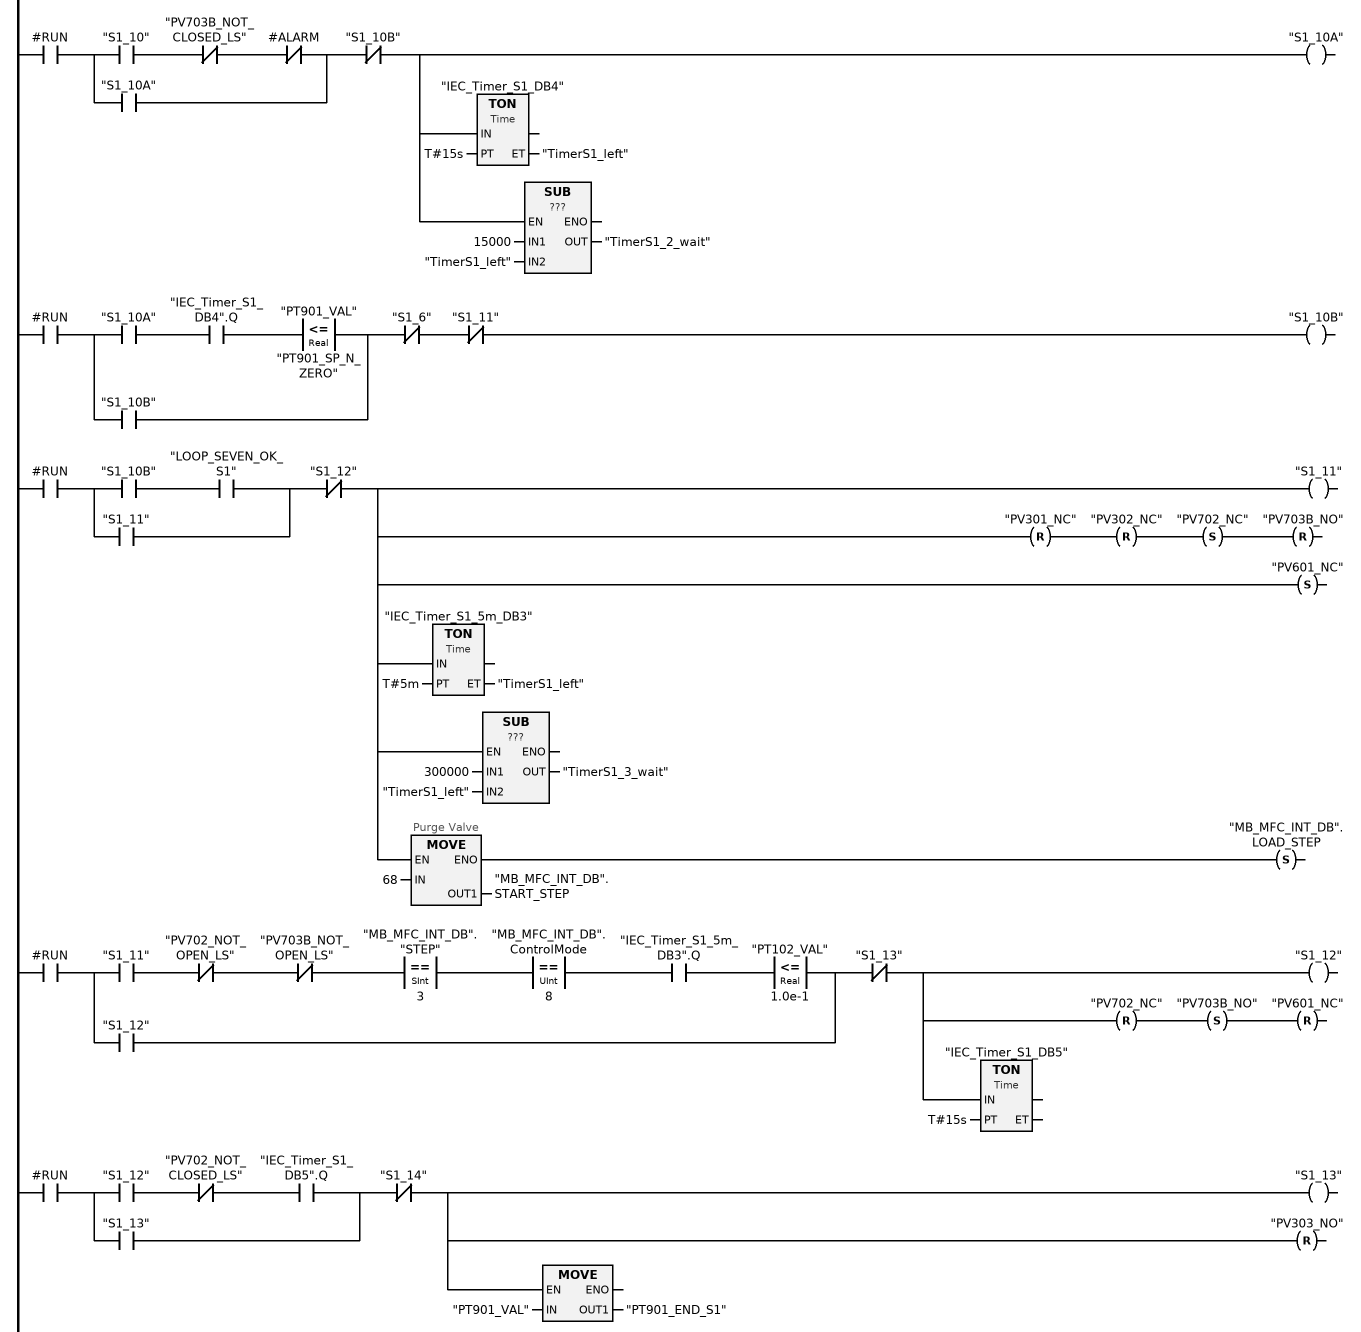
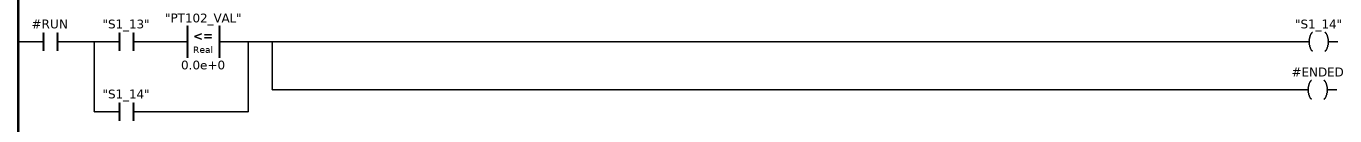
   "S1_0" := #RUN AND ((#START AND NOT #ALARM) OR "S1_0") AND NOT "S1_1";
   IF "S1_0" THEN
       "MB_MFC_INT_DB".MFC_MODE_SP := "MB_VAL_CONTROL_MODE_BUS";
       "MB_MFC_INT_DB".MFC_Setpoint := 0;
       "MB_MFC_INT_DB".START_STEP := 10;
       "MB_MFC_INT_DB".LOAD_STEP := TRUE;
       "MB_MFC_FLOAT_DB"."STEP" := -1;
   END_IF;
   "Timer_S1_DB_1S".TON(IN := "S1_0", PT := T#1S);
   IF "S1_0" THEN
       "GREEN_LIGHT" := FALSE;
       "YELLOW_LIGHT" := TRUE;
   END_IF;
   "S1_1" := #RUN AND (("S1_0" AND "Timer_S1_DB_1S".Q AND ("MB_MFC_INT_DB"."STEP" = 3) AND NOT #ALARM) OR "S1_1") AND NOT "S1_1A";
   IF "S1_1" THEN "PV703A_NO" := FALSE; END_IF;
   "S1_1A" := #RUN AND (("S1_1" AND NOT "PV703A_NOT_OPEN_LS" AND NOT #ALARM) OR "S1_1A") AND NOT "S1_2";
   IF "S1_1A" THEN
       "PV303_NO" := TRUE;
       "PV301_NC" := TRUE;
       "PV302_NC" := TRUE;
       "MB_MFC_INT_DB".MFC_Setpoint := "STEP1_MFC_FL_SP";
       "MB_MFC_INT_DB".START_STEP := 10;
       "MB_MFC_INT_DB".LOAD_STEP := TRUE;
   END_IF;
   "S1_2" := #RUN AND (("S1_1A" AND NOT #ALARM AND ("PT302_VAL" < "PT302_HIGH") AND ("MB_MFC_INT_DB"."STEP" = 3) AND ("MB_MFC_INT_DB".MFC_Setpoint = "STEP1_MFC_FL_SP")) OR "S1_2") AND NOT "S1_3";
   IF "S1_2" THEN "PV601_NC" := TRUE; END_IF;
   "S1_3" := #RUN AND (("S1_2" AND NOT #ALARM AND ("PT601_VAL" >= "PT302_CALC_90PRCT")) OR "S1_3") AND NOT "S1_4";
   IF "S1_3" THEN "PV702_NC" := TRUE; END_IF;
   "Timer_S1_DB_3S".TON(IN := "S1_3", PT := T#1.5s, ET => "TempDWord_A");
   "S1_4" := #RUN AND (("S1_3" AND "Timer_S1_DB_3S".Q AND NOT "PV702_NOT_OPEN_LS" AND NOT #ALARM) OR "S1_4") AND NOT "S1_5";
   IF "S1_4" THEN
       "PV601_NC" := FALSE;
       "PV702_NC" := FALSE;
   END_IF;
   "S1_5" := #RUN AND (("S1_4" AND NOT "PV702_NOT_CLOSED_LS" AND NOT #ALARM) OR "S1_5") AND NOT "S1_6";
   "IEC_Counter_S1_1".CTU(CU := "S1_7", R := "S1_2", PV := "STEP1_LOOPS", CV => "Counter_S1");
   "LOOP_SEVEN_OK_S1" := "IEC_Counter_S1_1".Q;
   "S1_6" := #RUN AND ((("S1_5" OR ("S1_10B" AND NOT "LOOP_SEVEN_OK_S1")) AND NOT #ALARM) OR "S1_6") AND NOT "S1_7";
   IF "S1_6" THEN
       "PV701_NC" := TRUE;
       "PT901_SAVE" := "PT901_VAL" - 1.0;
   END_IF;
   IF "S1_6" AND ("PT601_VAL" < 3.5) THEN "PV601_NC" := TRUE; END_IF;
   "S1_7" := #RUN AND (("S1_6" AND NOT "PV701_NOT_OPEN_LS" AND ("PT901_VAL" >= "PT901_SP_N")) OR "S1_7") AND NOT "S1_7A";
   IF "S1_7" THEN
       "PV701_NC" := FALSE;
       "PV601_NC" := FALSE;
   END_IF;
   "S1_7A" := #RUN AND (("S1_7" AND NOT "PV701_NOT_CLOSED_LS" AND "Timer_S1_DB_5S".Q AND ("PT901_VAL" >= "PT901_SAVE")) OR "S1_7A") AND NOT "S1_8";
   "S1_8" := #RUN AND (("S1_7A" AND NOT #ALARM) OR "S1_8") AND NOT "S1_9";
   IF "S1_8" THEN "PV703B_NO" := FALSE; END_IF;
   "S1_9" := #RUN AND (("S1_8" AND NOT "PV703B_NOT_OPEN_LS" AND ("PT901_VAL" <= "PT901_SP_PV703B_OPEN") AND NOT #ALARM) OR "S1_9") AND NOT "S1_10";
   "IEC_Timer_S1_DB3".TON(IN := "S1_9", PT := T#150s, ET => "TimerS1_left");
   IF "S1_9" THEN "TimerS1_1_wait" := 150000 - "TimerS1_left"; END_IF;
   "S1_10" := #RUN AND (("S1_9" AND "IEC_Timer_S1_DB3".Q AND ("PT901_VAL" <= 0.2)) OR "S1_10") AND NOT "S1_10A";
   IF "S1_10" THEN "PV703B_NO" := TRUE; END_IF;
   "S1_10A" := #RUN AND (("S1_10" AND NOT "PV703B_NOT_CLOSED_LS" AND NOT #ALARM) OR "S1_10A") AND NOT "S1_10B";
   "IEC_Timer_S1_DB4".TON(IN := "S1_10A", PT := T#15s, ET => "TimerS1_left");
   IF "S1_10A" THEN "TimerS1_2_wait" := 15000 - "TimerS1_left"; END_IF;
   "S1_10B" := #RUN AND (("S1_10A" AND "IEC_Timer_S1_DB4".Q AND ("PT901_VAL" <= "PT901_SP_N_ZERO")) OR "S1_10B") AND NOT "S1_6" AND NOT "S1_11";
   "S1_11" := #RUN AND (("S1_10B" AND "LOOP_SEVEN_OK_S1") OR "S1_11") AND NOT "S1_12";
   IF "S1_11" THEN
       "PV301_NC" := FALSE;
       "PV302_NC" := FALSE;
       "PV702_NC" := TRUE;
       "PV703B_NO" := FALSE;
       "PV601_NC" := TRUE;
   END_IF;
   "IEC_Timer_S1_5m_DB3".TON(IN := "S1_11", PT := T#5m, ET => "TimerS1_left");
   IF "S1_11" THEN
       "TimerS1_3_wait" := 300000 - "TimerS1_left";
       "MB_MFC_INT_DB".START_STEP := 68;   // Purge Valve
       "MB_MFC_INT_DB".LOAD_STEP := TRUE;
   END_IF;
   "S1_12" := #RUN AND (("S1_11" AND NOT "PV702_NOT_OPEN_LS" AND NOT "PV703B_NOT_OPEN_LS" AND ("MB_MFC_INT_DB"."STEP" = 3) AND ("MB_MFC_INT_DB".ControlMode = 8) AND "IEC_Timer_S1_5m_DB3".Q AND ("PT102_VAL" <= 1.0e-1)) OR "S1_12") AND NOT "S1_13";
   IF "S1_12" THEN
       "PV702_NC" := FALSE;
       "PV703B_NO" := TRUE;
       "PV601_NC" := FALSE;
   END_IF;
   "IEC_Timer_S1_DB5".TON(IN := "S1_12", PT := T#15s);
   "S1_13" := #RUN AND (("S1_12" AND NOT "PV702_NOT_CLOSED_LS" AND "IEC_Timer_S1_DB5".Q) OR "S1_13") AND NOT "S1_14";
   IF "S1_13" THEN
       "PV303_NO" := FALSE;
       "PT901_END_S1" := "PT901_VAL";
   END_IF;
   "S1_14" := #RUN AND (("S1_13" AND ("PT102_VAL" <= 0.0e+0)) OR "S1_14");
   #ENDED := "S1_14";
END_REGION

REGION Network 4
   // Timers
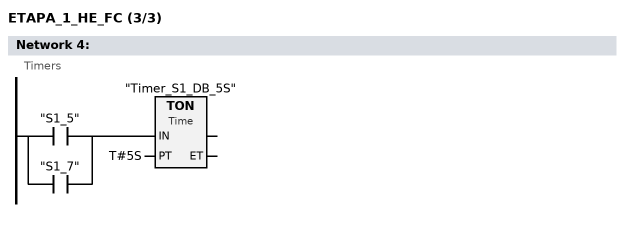
   "Timer_S1_DB_5S".TON(IN := "S1_5" OR "S1_7", PT := T#5S);
END_REGION
END_FUNCTION

FUNCTION "MB_READ_MX" : Void   // FC23, LAD
{ S7_Optimized_Access := 'FALSE' }
VERSION : 0.1
   VAR_TEMP   // added for the SCL form of the ladder/FBD networks
      _w1 : Bool;
      _w2 : Bool;
   END_VAR
BEGIN

REGION Network 1
   // MODBUS MASTER Cyclic Read
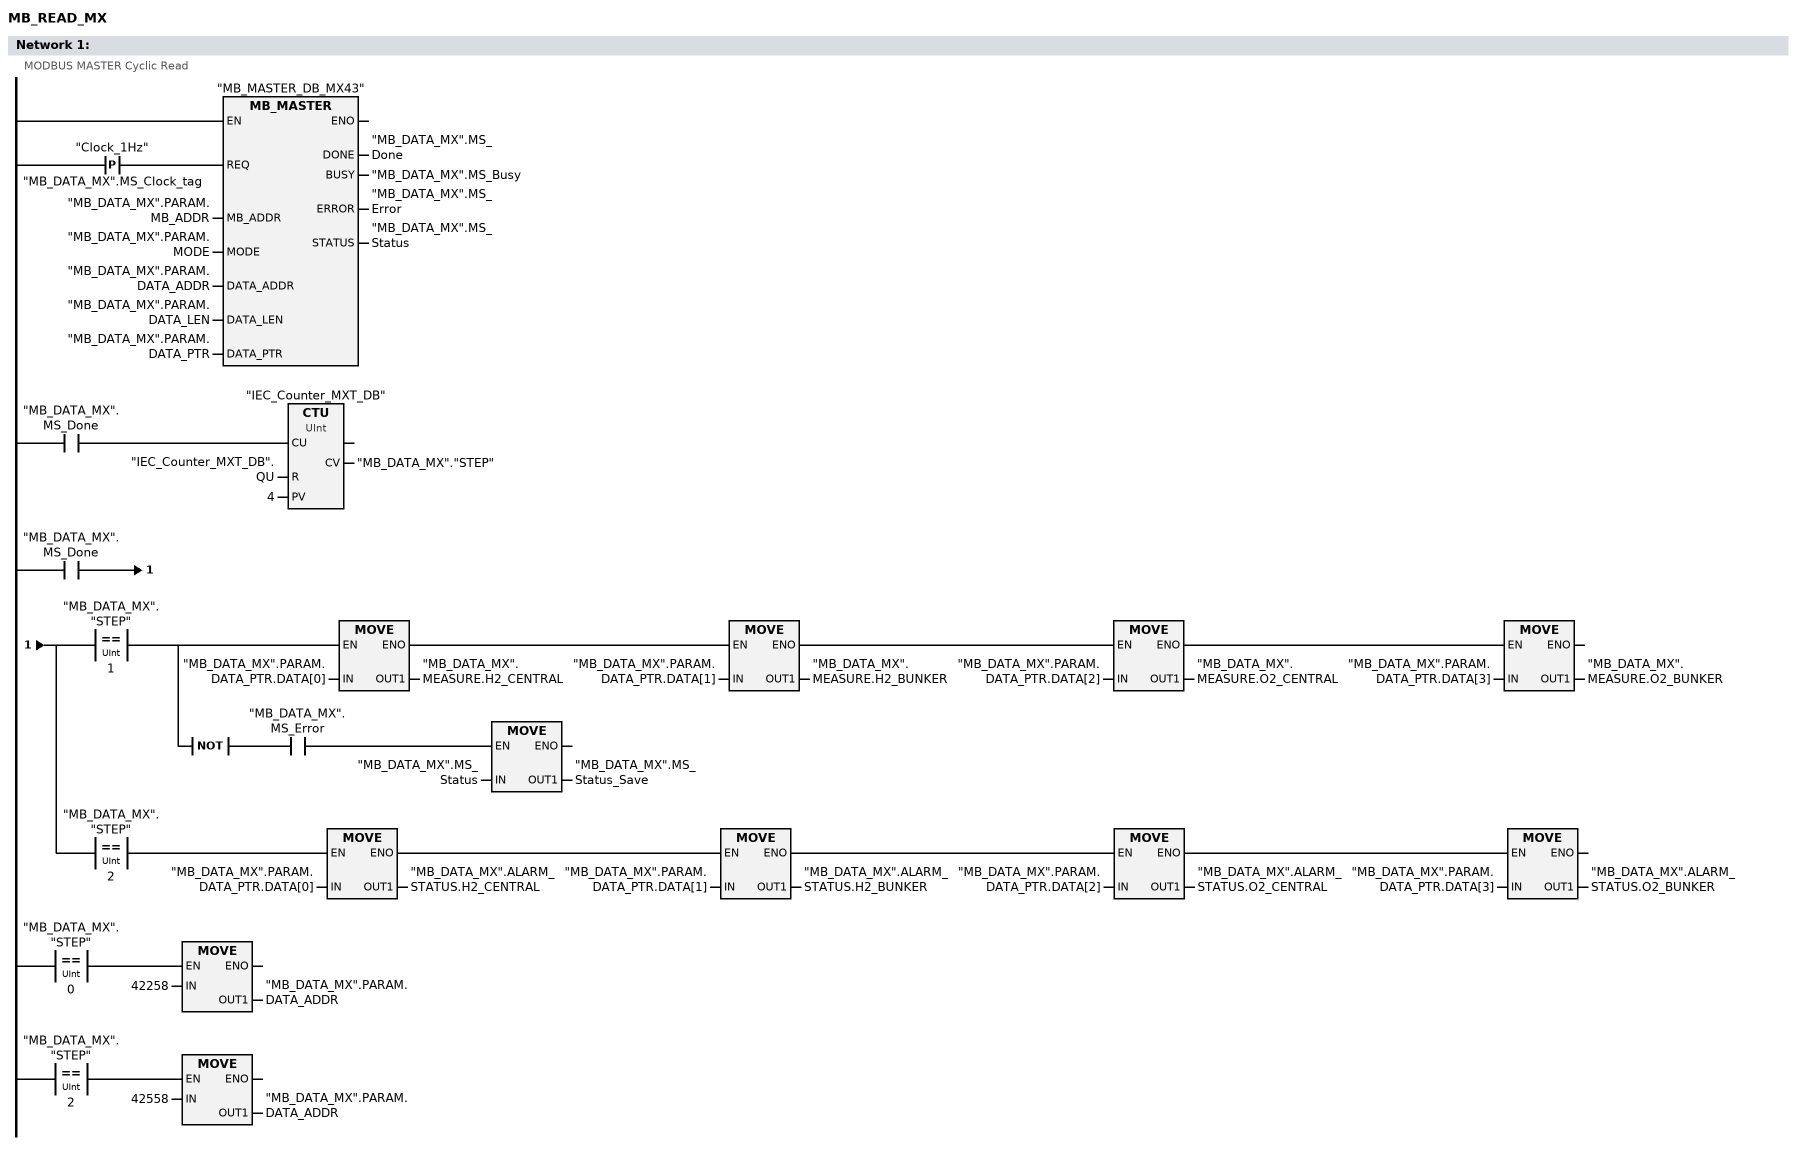
   #_w1 := "Clock_1Hz" AND NOT "MB_DATA_MX".MS_Clock_tag;   // rising edge of "Clock_1Hz"
   "MB_DATA_MX".MS_Clock_tag := "Clock_1Hz";
   "MB_MASTER_DB_MX43"(REQ := #_w1,   // MB_MASTER
                       MB_ADDR := "MB_DATA_MX".PARAM.MB_ADDR,
                       MODE := "MB_DATA_MX".PARAM.MODE,
                       DATA_ADDR := "MB_DATA_MX".PARAM.DATA_ADDR,
                       DATA_LEN := "MB_DATA_MX".PARAM.DATA_LEN,
                       DATA_PTR := "MB_DATA_MX".PARAM.DATA_PTR,
                       DONE => "MB_DATA_MX".MS_Done,
                       BUSY => "MB_DATA_MX".MS_Busy,
                       ERROR => "MB_DATA_MX".MS_Error,
                       STATUS => "MB_DATA_MX".MS_Status);
   "IEC_Counter_MXT_DB".CTU(CU := "MB_DATA_MX".MS_Done,
                           R := "IEC_Counter_MXT_DB".QU,
                           PV := 4,
                           CV => "MB_DATA_MX"."STEP");
   #_w2 := "MB_DATA_MX".MS_Done AND ("MB_DATA_MX"."STEP" = 1);
   IF #_w2 THEN
       "MB_DATA_MX".MEASURE.H2_CENTRAL := "MB_DATA_MX".PARAM.DATA_PTR.DATA[0];
       "MB_DATA_MX".MEASURE.H2_BUNKER := "MB_DATA_MX".PARAM.DATA_PTR.DATA[1];
       "MB_DATA_MX".MEASURE.O2_CENTRAL := "MB_DATA_MX".PARAM.DATA_PTR.DATA[2];
       "MB_DATA_MX".MEASURE.O2_BUNKER := "MB_DATA_MX".PARAM.DATA_PTR.DATA[3];
   END_IF;
   IF NOT #_w2 AND "MB_DATA_MX".MS_Error THEN "MB_DATA_MX".MS_Status_Save := "MB_DATA_MX".MS_Status; END_IF;
   IF "MB_DATA_MX".MS_Done AND ("MB_DATA_MX"."STEP" = 2) THEN
       "MB_DATA_MX".ALARM_STATUS.H2_CENTRAL := "MB_DATA_MX".PARAM.DATA_PTR.DATA[0];
       "MB_DATA_MX".ALARM_STATUS.H2_BUNKER := "MB_DATA_MX".PARAM.DATA_PTR.DATA[1];
       "MB_DATA_MX".ALARM_STATUS.O2_CENTRAL := "MB_DATA_MX".PARAM.DATA_PTR.DATA[2];
       "MB_DATA_MX".ALARM_STATUS.O2_BUNKER := "MB_DATA_MX".PARAM.DATA_PTR.DATA[3];
   END_IF;
   IF "MB_DATA_MX"."STEP" = 0 THEN "MB_DATA_MX".PARAM.DATA_ADDR := 42258; END_IF;
   IF "MB_DATA_MX"."STEP" = 2 THEN "MB_DATA_MX".PARAM.DATA_ADDR := 42558; END_IF;
END_REGION
END_FUNCTION

ORGANIZATION_BLOCK "Main"   // OB1, LAD, ProgramCycle
TITLE = "Main Program Sweep (Cycle)"
{ S7_Optimized_Access := 'FALSE' }
VERSION : 0.1
// Main with He Purging, Step 2 is Bypassed
   VAR_TEMP   // added for the SCL form of the ladder/FBD networks
      _w1 : Bool;
   END_VAR
BEGIN

REGION Network 1
   // TOP LOGIC
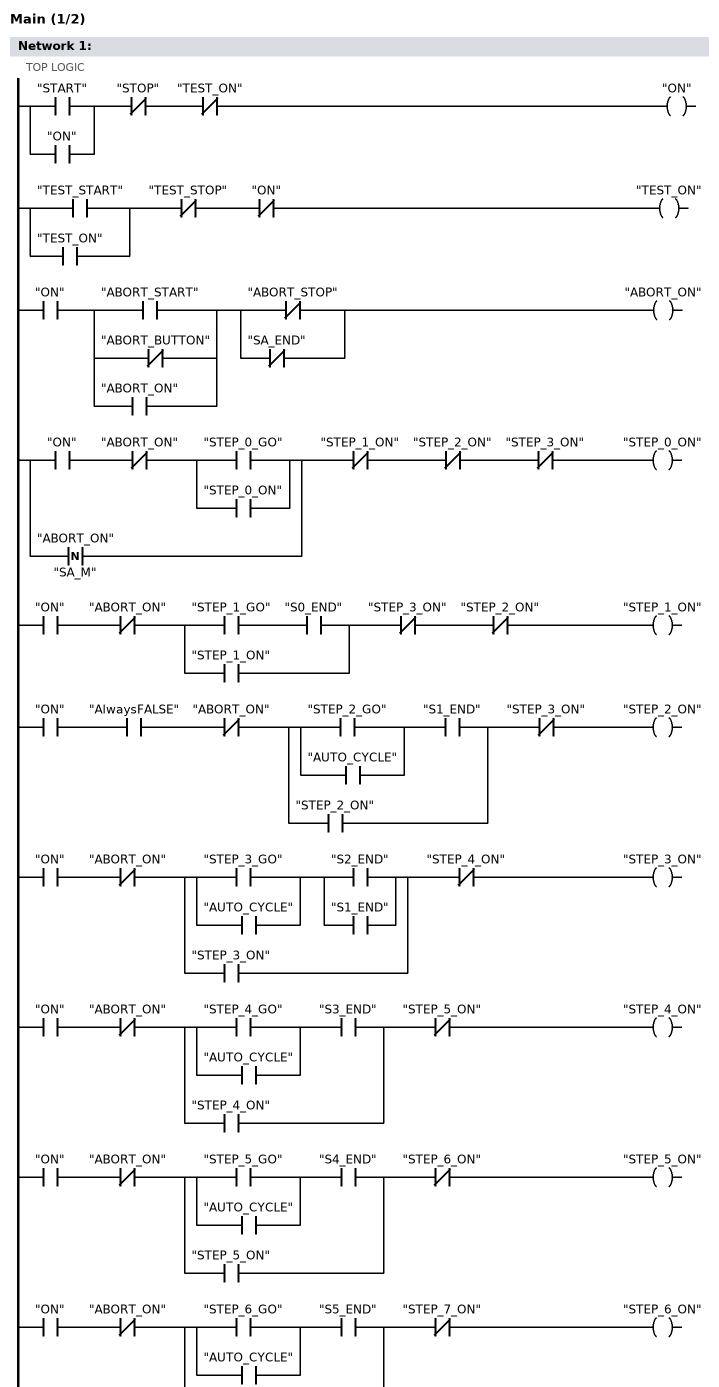
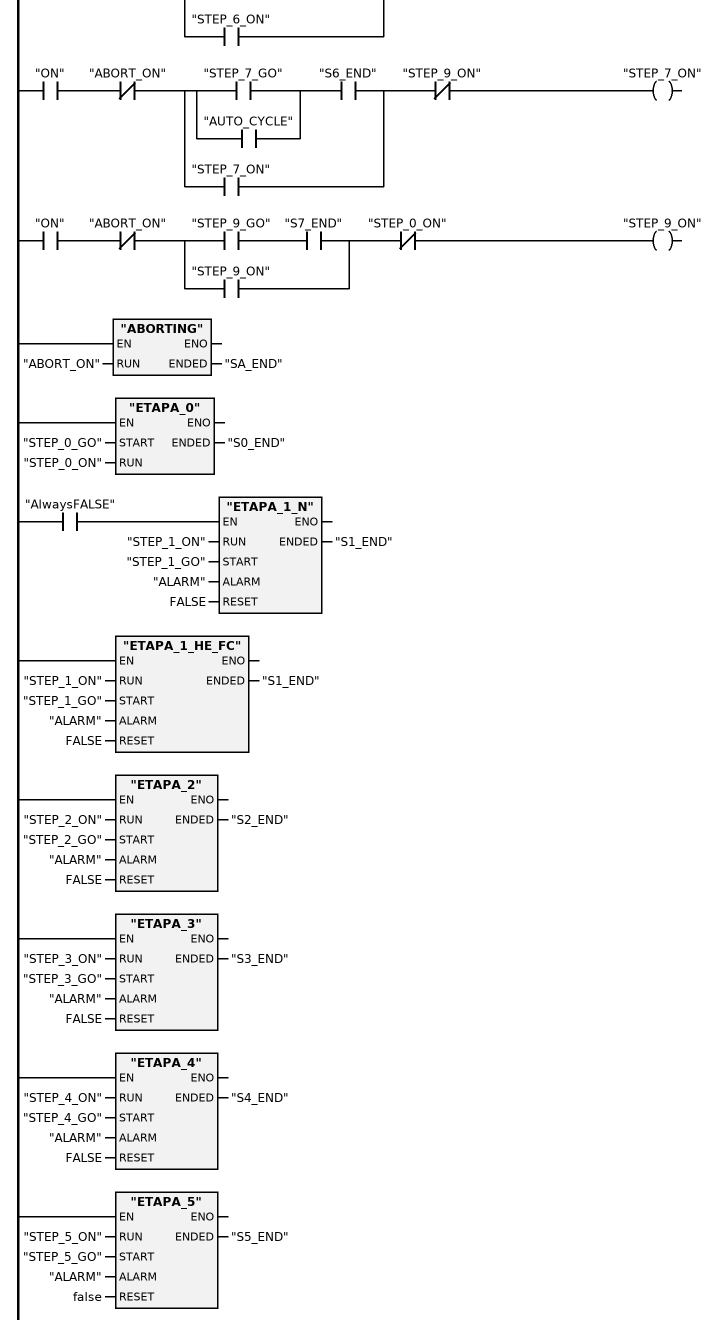
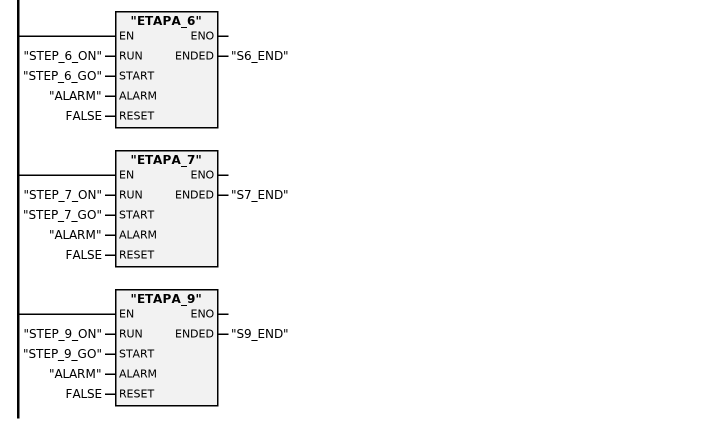
   RUNG wire#powerrail
      Contact( "START" )
      wire#w1
      I_Contact( "STOP" )
      I_Contact( "TEST_ON" )
      Coil( "ON" )
   END_RUNG
   RUNG wire#powerrail
      Contact( "ON" )
   END_RUNG wire#w1
   RUNG wire#powerrail
      Contact( "TEST_START" )
      wire#w2
      I_Contact( "TEST_STOP" )
      I_Contact( "ON" )
      Coil( "TEST_ON" )
   END_RUNG
   RUNG wire#powerrail
      Contact( "TEST_ON" )
   END_RUNG wire#w2
   RUNG wire#powerrail
      Contact( "ON" )
      wire#w3
      Contact( "ABORT_START" )
      wire#w4
      I_Contact( "ABORT_STOP" )
      wire#w5
      Coil( "ABORT_ON" )
   END_RUNG
   RUNG wire#w3
      I_Contact( "ABORT_BUTTON" )
   END_RUNG wire#w4
   RUNG wire#w3
      Contact( "ABORT_ON" )
   END_RUNG wire#w4
   RUNG wire#w4
      I_Contact( "SA_END" )
   END_RUNG wire#w5
   RUNG wire#powerrail
      Contact( "ON" )
      I_Contact( "ABORT_ON" )
      wire#w6
      Contact( "STEP_0_GO" )
      wire#w7
      I_Contact( "STEP_1_ON" )
      I_Contact( "STEP_2_ON" )
      I_Contact( "STEP_3_ON" )
      Coil( "STEP_0_ON" )
   END_RUNG
   RUNG wire#w6
      Contact( "STEP_0_ON" )
   END_RUNG wire#w7
   RUNG wire#powerrail
      N_Contact(operand := "ABORT_ON", bit := "SA_M")
   END_RUNG wire#w7
   RUNG wire#powerrail
      Contact( "ON" )
      I_Contact( "ABORT_ON" )
      wire#w8
      Contact( "STEP_1_GO" )
      Contact( "S0_END" )
      wire#w9
      I_Contact( "STEP_3_ON" )
      I_Contact( "STEP_2_ON" )
      Coil( "STEP_1_ON" )
   END_RUNG
   RUNG wire#w8
      Contact( "STEP_1_ON" )
   END_RUNG wire#w9
   RUNG wire#powerrail
      Contact( "ON" )
      Contact( "AlwaysFALSE" )
      I_Contact( "ABORT_ON" )
      wire#w10
      Contact( "STEP_2_GO" )
      wire#w11
      Contact( "S1_END" )
      wire#w12
      I_Contact( "STEP_3_ON" )
      Coil( "STEP_2_ON" )
   END_RUNG
   RUNG wire#w10
      Contact( "AUTO_CYCLE" )
   END_RUNG wire#w11
   RUNG wire#w10
      Contact( "STEP_2_ON" )
   END_RUNG wire#w12
   RUNG wire#powerrail
      Contact( "ON" )
      I_Contact( "ABORT_ON" )
      wire#w13
      Contact( "STEP_3_GO" )
      wire#w14
      Contact( "S2_END" )
      wire#w15
      I_Contact( "STEP_4_ON" )
      Coil( "STEP_3_ON" )
   END_RUNG
   RUNG wire#w13
      Contact( "AUTO_CYCLE" )
   END_RUNG wire#w14
   RUNG wire#w14
      Contact( "S1_END" )
   END_RUNG wire#w15
   RUNG wire#w13
      Contact( "STEP_3_ON" )
   END_RUNG wire#w15
   RUNG wire#powerrail
      Contact( "ON" )
      I_Contact( "ABORT_ON" )
      wire#w16
      Contact( "STEP_4_GO" )
      wire#w17
      Contact( "S3_END" )
      wire#w18
      I_Contact( "STEP_5_ON" )
      Coil( "STEP_4_ON" )
   END_RUNG
   RUNG wire#w16
      Contact( "AUTO_CYCLE" )
   END_RUNG wire#w17
   RUNG wire#w16
      Contact( "STEP_4_ON" )
   END_RUNG wire#w18
   RUNG wire#powerrail
      Contact( "ON" )
      I_Contact( "ABORT_ON" )
      wire#w19
      Contact( "STEP_5_GO" )
      wire#w20
      Contact( "S4_END" )
      wire#w21
      I_Contact( "STEP_6_ON" )
      Coil( "STEP_5_ON" )
   END_RUNG
   RUNG wire#w19
      Contact( "AUTO_CYCLE" )
   END_RUNG wire#w20
   RUNG wire#w19
      Contact( "STEP_5_ON" )
   END_RUNG wire#w21
   RUNG wire#powerrail
      Contact( "ON" )
      I_Contact( "ABORT_ON" )
      wire#w22
      Contact( "STEP_6_GO" )
      wire#w23
      Contact( "S5_END" )
      wire#w24
      I_Contact( "STEP_7_ON" )
      Coil( "STEP_6_ON" )
   END_RUNG
   RUNG wire#w22
      Contact( "AUTO_CYCLE" )
   END_RUNG wire#w23
   RUNG wire#w22
      Contact( "STEP_6_ON" )
   END_RUNG wire#w24
   RUNG wire#powerrail
      Contact( "ON" )
      I_Contact( "ABORT_ON" )
      wire#w25
      Contact( "STEP_7_GO" )
      wire#w26
      Contact( "S6_END" )
      wire#w27
      I_Contact( "STEP_9_ON" )
      Coil( "STEP_7_ON" )
   END_RUNG
   RUNG wire#w25
      Contact( "AUTO_CYCLE" )
   END_RUNG wire#w26
   RUNG wire#w25
      Contact( "STEP_7_ON" )
   END_RUNG wire#w27
   RUNG wire#powerrail
      Contact( "ON" )
      I_Contact( "ABORT_ON" )
      wire#w28
      Contact( "STEP_9_GO" )
      Contact( "S7_END" )
      wire#w29
      I_Contact( "STEP_0_ON" )
      Coil( "STEP_9_ON" )
   END_RUNG
   RUNG wire#w28
      Contact( "STEP_9_ON" )
   END_RUNG wire#w29
   RUNG wire#powerrail
      "ABORTING"(RUN := "ABORT_ON", ENDED => "SA_END")
   END_RUNG
   RUNG wire#powerrail
      "ETAPA_0"(START := "STEP_0_GO", RUN := "STEP_0_ON", ENDED => "S0_END")
   END_RUNG
   RUNG wire#powerrail
      Contact( "AlwaysFALSE" )
      "ETAPA_1_N"(RUN := "STEP_1_ON", START := "STEP_1_GO", ALARM := "ALARM", RESET := FALSE, ENDED => "S1_END")
   END_RUNG
   RUNG wire#powerrail
      "ETAPA_1_HE_FC"(RUN := "STEP_1_ON", START := "STEP_1_GO", ALARM := "ALARM", RESET := FALSE, ENDED => "S1_END")
   END_RUNG
   RUNG wire#powerrail
      "ETAPA_2"(RUN := "STEP_2_ON", START := "STEP_2_GO", ALARM := "ALARM", RESET := FALSE, ENDED => "S2_END")
   END_RUNG
   RUNG wire#powerrail
      "ETAPA_3"(RUN := "STEP_3_ON", START := "STEP_3_GO", ALARM := "ALARM", RESET := FALSE, ENDED => "S3_END")
   END_RUNG
   RUNG wire#powerrail
      "ETAPA_4"(RUN := "STEP_4_ON", START := "STEP_4_GO", ALARM := "ALARM", RESET := FALSE, ENDED => "S4_END")
   END_RUNG
   RUNG wire#powerrail
      "ETAPA_5"(RUN := "STEP_5_ON", START := "STEP_5_GO", ALARM := "ALARM", RESET := false, ENDED => "S5_END")
   END_RUNG
   RUNG wire#powerrail
      "ETAPA_6"(RUN := "STEP_6_ON", START := "STEP_6_GO", ALARM := "ALARM", RESET := FALSE, ENDED => "S6_END")
   END_RUNG
   RUNG wire#powerrail
      "ETAPA_7"(RUN := "STEP_7_ON", START := "STEP_7_GO", ALARM := "ALARM", RESET := FALSE, ENDED => "S7_END")
   END_RUNG
   RUNG wire#powerrail
      "ETAPA_9"(RUN := "STEP_9_ON", START := "STEP_9_GO", ALARM := "ALARM", RESET := FALSE, ENDED => "S9_END")
   END_RUNG
   // the same network as SCL:
   "ON" := ("START" OR "ON") AND NOT "STOP" AND NOT "TEST_ON";
   "TEST_ON" := ("TEST_START" OR "TEST_ON") AND NOT "TEST_STOP" AND NOT "ON";
   "ABORT_ON" := "ON" AND ("ABORT_START" OR NOT "ABORT_BUTTON" OR "ABORT_ON") AND (NOT "ABORT_STOP" OR NOT "SA_END");
   #_w1 := NOT "ABORT_ON" AND "SA_M";   // falling edge of "ABORT_ON"
   "SA_M" := "ABORT_ON";
   "STEP_0_ON" := (("ON" AND NOT "ABORT_ON" AND ("STEP_0_GO" OR "STEP_0_ON")) OR #_w1) AND NOT "STEP_1_ON" AND NOT "STEP_2_ON" AND NOT "STEP_3_ON";
   "STEP_1_ON" := "ON" AND NOT "ABORT_ON" AND (("STEP_1_GO" AND "S0_END") OR "STEP_1_ON") AND NOT "STEP_3_ON" AND NOT "STEP_2_ON";
   "STEP_2_ON" := "ON" AND "AlwaysFALSE" AND NOT "ABORT_ON" AND ((("STEP_2_GO" OR "AUTO_CYCLE") AND "S1_END") OR "STEP_2_ON") AND NOT "STEP_3_ON";
   "STEP_3_ON" := "ON" AND NOT "ABORT_ON" AND ((("STEP_3_GO" OR "AUTO_CYCLE") AND ("S2_END" OR "S1_END")) OR "STEP_3_ON") AND NOT "STEP_4_ON";
   "STEP_4_ON" := "ON" AND NOT "ABORT_ON" AND ((("STEP_4_GO" OR "AUTO_CYCLE") AND "S3_END") OR "STEP_4_ON") AND NOT "STEP_5_ON";
   "STEP_5_ON" := "ON" AND NOT "ABORT_ON" AND ((("STEP_5_GO" OR "AUTO_CYCLE") AND "S4_END") OR "STEP_5_ON") AND NOT "STEP_6_ON";
   "STEP_6_ON" := "ON" AND NOT "ABORT_ON" AND ((("STEP_6_GO" OR "AUTO_CYCLE") AND "S5_END") OR "STEP_6_ON") AND NOT "STEP_7_ON";
   "STEP_7_ON" := "ON" AND NOT "ABORT_ON" AND ((("STEP_7_GO" OR "AUTO_CYCLE") AND "S6_END") OR "STEP_7_ON") AND NOT "STEP_9_ON";
   "STEP_9_ON" := "ON" AND NOT "ABORT_ON" AND (("STEP_9_GO" AND "S7_END") OR "STEP_9_ON") AND NOT "STEP_0_ON";
   "ABORTING"(RUN := "ABORT_ON", ENDED => "SA_END");
   "ETAPA_0"(START := "STEP_0_GO", RUN := "STEP_0_ON", ENDED => "S0_END");
   IF "AlwaysFALSE" THEN
       "ETAPA_1_N"(RUN := "STEP_1_ON", START := "STEP_1_GO", ALARM := "ALARM", RESET := FALSE, ENDED => "S1_END");
   END_IF;
   "ETAPA_1_HE_FC"(RUN := "STEP_1_ON",
                   START := "STEP_1_GO",
                   ALARM := "ALARM",
                   RESET := FALSE,
                   ENDED => "S1_END");
   "ETAPA_2"(RUN := "STEP_2_ON", START := "STEP_2_GO", ALARM := "ALARM", RESET := FALSE, ENDED => "S2_END");
   "ETAPA_3"(RUN := "STEP_3_ON", START := "STEP_3_GO", ALARM := "ALARM", RESET := FALSE, ENDED => "S3_END");
   "ETAPA_4"(RUN := "STEP_4_ON", START := "STEP_4_GO", ALARM := "ALARM", RESET := FALSE, ENDED => "S4_END");
   "ETAPA_5"(RUN := "STEP_5_ON", START := "STEP_5_GO", ALARM := "ALARM", RESET := false, ENDED => "S5_END");
   "ETAPA_6"(RUN := "STEP_6_ON", START := "STEP_6_GO", ALARM := "ALARM", RESET := FALSE, ENDED => "S6_END");
   "ETAPA_7"(RUN := "STEP_7_ON", START := "STEP_7_GO", ALARM := "ALARM", RESET := FALSE, ENDED => "S7_END");
   "ETAPA_9"(RUN := "STEP_9_ON", START := "STEP_9_GO", ALARM := "ALARM", RESET := FALSE, ENDED => "S9_END");
END_REGION

REGION Network 2
   // ALARM Block
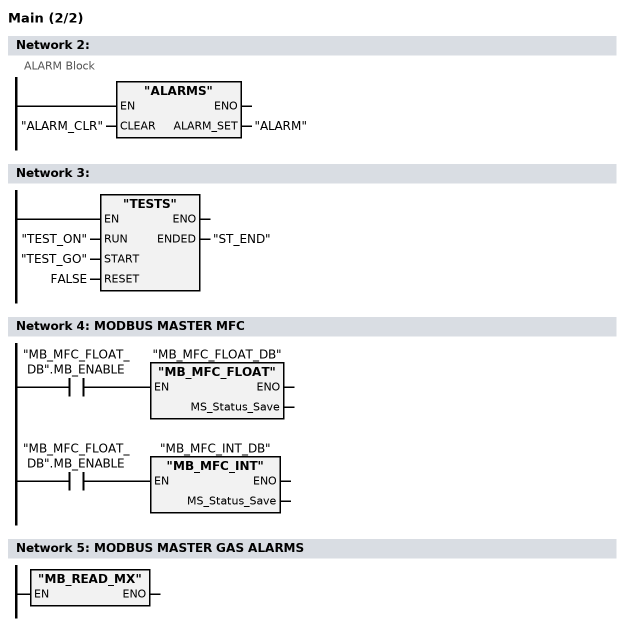
   RUNG wire#powerrail
      "ALARMS"(CLEAR := "ALARM_CLR", ALARM_SET => "ALARM")
   END_RUNG
   // the same network as SCL:
   "ALARMS"(CLEAR := "ALARM_CLR", ALARM_SET => "ALARM");
END_REGION

REGION Network 3
   RUNG wire#powerrail
      "TESTS"(RUN := "TEST_ON", START := "TEST_GO", RESET := FALSE, ENDED => "ST_END")
   END_RUNG
   // the same network as SCL:
   "TESTS"(RUN := "TEST_ON", START := "TEST_GO", RESET := FALSE, ENDED => "ST_END");
END_REGION

REGION Network 4: MODBUS MASTER MFC
   RUNG wire#powerrail
      Contact( "MB_MFC_FLOAT_DB".MB_ENABLE )
      "MB_MFC_FLOAT_DB"(MS_Status_Save =>)
   END_RUNG
   RUNG wire#powerrail
      Contact( "MB_MFC_FLOAT_DB".MB_ENABLE )
      "MB_MFC_INT_DB"(MS_Status_Save =>)
   END_RUNG
   // the same network as SCL:
   IF "MB_MFC_FLOAT_DB".MB_ENABLE THEN
       "MB_MFC_FLOAT_DB"();   // "MB_MFC_FLOAT"
   END_IF;
   IF "MB_MFC_FLOAT_DB".MB_ENABLE THEN
       "MB_MFC_INT_DB"();   // "MB_MFC_INT"
   END_IF;
END_REGION

REGION Network 5: MODBUS MASTER GAS ALARMS
   RUNG wire#powerrail
      "MB_READ_MX"()
   END_RUNG
   // the same network as SCL:
   "MB_READ_MX"();
END_REGION
END_ORGANIZATION_BLOCK

ORGANIZATION_BLOCK "PV_Cyclic interrupt"   // OB30, LAD, CyclicInterrupt
{ S7_Optimized_Access := 'FALSE' }
VERSION : 0.1
BEGIN

REGION Network 1
   // Calculations
END_REGION

REGION Network 2
   // ABORTING
END_REGION

REGION Network 3
   // Analog Input Scaling Module AI_1
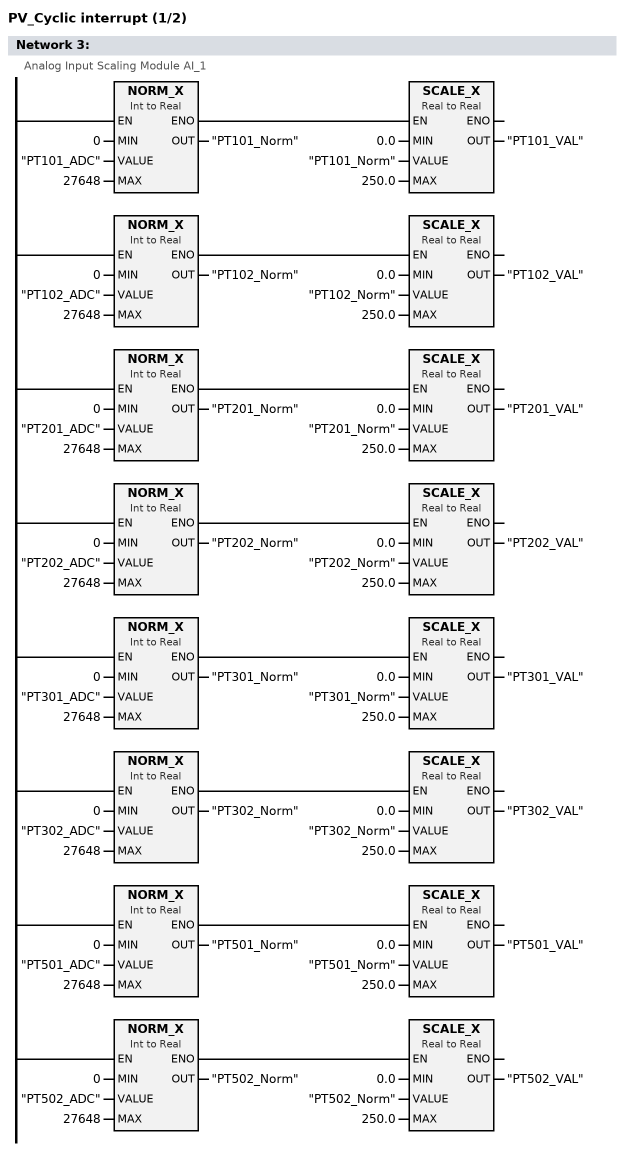
   RUNG wire#powerrail
      { S7_Templates := "[SrcType := Int, DestType := Real]" } Normalize(min := 0, value := "PT101_ADC", max := 27648, out => "PT101_Norm")
      { S7_Templates := "[SrcType := Real, DestType := Real]" } Scale(min := 0.0, value := "PT101_Norm", max := 250.0, out => "PT101_VAL")
   END_RUNG
   RUNG wire#powerrail
      { S7_Templates := "[SrcType := Int, DestType := Real]" } Normalize(min := 0, value := "PT102_ADC", max := 27648, out => "PT102_Norm")
      { S7_Templates := "[SrcType := Real, DestType := Real]" } Scale(min := 0.0, value := "PT102_Norm", max := 250.0, out => "PT102_VAL")
   END_RUNG
   RUNG wire#powerrail
      { S7_Templates := "[SrcType := Int, DestType := Real]" } Normalize(min := 0, value := "PT201_ADC", max := 27648, out => "PT201_Norm")
      { S7_Templates := "[SrcType := Real, DestType := Real]" } Scale(min := 0.0, value := "PT201_Norm", max := 250.0, out => "PT201_VAL")
   END_RUNG
   RUNG wire#powerrail
      { S7_Templates := "[SrcType := Int, DestType := Real]" } Normalize(min := 0, value := "PT202_ADC", max := 27648, out => "PT202_Norm")
      { S7_Templates := "[SrcType := Real, DestType := Real]" } Scale(min := 0.0, value := "PT202_Norm", max := 250.0, out => "PT202_VAL")
   END_RUNG
   RUNG wire#powerrail
      { S7_Templates := "[SrcType := Int, DestType := Real]" } Normalize(min := 0, value := "PT301_ADC", max := 27648, out => "PT301_Norm")
      { S7_Templates := "[SrcType := Real, DestType := Real]" } Scale(min := 0.0, value := "PT301_Norm", max := 250.0, out => "PT301_VAL")
   END_RUNG
   RUNG wire#powerrail
      { S7_Templates := "[SrcType := Int, DestType := Real]" } Normalize(min := 0, value := "PT302_ADC", max := 27648, out => "PT302_Norm")
      { S7_Templates := "[SrcType := Real, DestType := Real]" } Scale(min := 0.0, value := "PT302_Norm", max := 250.0, out => "PT302_VAL")
   END_RUNG
   RUNG wire#powerrail
      { S7_Templates := "[SrcType := Int, DestType := Real]" } Normalize(min := 0, value := "PT501_ADC", max := 27648, out => "PT501_Norm")
      { S7_Templates := "[SrcType := Real, DestType := Real]" } Scale(min := 0.0, value := "PT501_Norm", max := 250.0, out => "PT501_VAL")
   END_RUNG
   RUNG wire#powerrail
      { S7_Templates := "[SrcType := Int, DestType := Real]" } Normalize(min := 0, value := "PT502_ADC", max := 27648, out => "PT502_Norm")
      { S7_Templates := "[SrcType := Real, DestType := Real]" } Scale(min := 0.0, value := "PT502_Norm", max := 250.0, out => "PT502_VAL")
   END_RUNG
   // the same network as SCL:
   "PT101_Norm" := NORM_X(MIN := 0, VALUE := "PT101_ADC", MAX := 27648);
   "PT101_VAL" := SCALE_X(MIN := 0.0, VALUE := "PT101_Norm", MAX := 250.0);
   "PT102_Norm" := NORM_X(MIN := 0, VALUE := "PT102_ADC", MAX := 27648);
   "PT102_VAL" := SCALE_X(MIN := 0.0, VALUE := "PT102_Norm", MAX := 250.0);
   "PT201_Norm" := NORM_X(MIN := 0, VALUE := "PT201_ADC", MAX := 27648);
   "PT201_VAL" := SCALE_X(MIN := 0.0, VALUE := "PT201_Norm", MAX := 250.0);
   "PT202_Norm" := NORM_X(MIN := 0, VALUE := "PT202_ADC", MAX := 27648);
   "PT202_VAL" := SCALE_X(MIN := 0.0, VALUE := "PT202_Norm", MAX := 250.0);
   "PT301_Norm" := NORM_X(MIN := 0, VALUE := "PT301_ADC", MAX := 27648);
   "PT301_VAL" := SCALE_X(MIN := 0.0, VALUE := "PT301_Norm", MAX := 250.0);
   "PT302_Norm" := NORM_X(MIN := 0, VALUE := "PT302_ADC", MAX := 27648);
   "PT302_VAL" := SCALE_X(MIN := 0.0, VALUE := "PT302_Norm", MAX := 250.0);
   "PT501_Norm" := NORM_X(MIN := 0, VALUE := "PT501_ADC", MAX := 27648);
   "PT501_VAL" := SCALE_X(MIN := 0.0, VALUE := "PT501_Norm", MAX := 250.0);
   "PT502_Norm" := NORM_X(MIN := 0, VALUE := "PT502_ADC", MAX := 27648);
   "PT502_VAL" := SCALE_X(MIN := 0.0, VALUE := "PT502_Norm", MAX := 250.0);
END_REGION

REGION Network 4
   // Analog Input Scaling Module AI_2
